(* Logix 5000 project; controller MV vendor 1 type 14 code 217 rev 31.11; software revision 31.00; part 32 of 53 *)
(* tags used below, declared in another part *)
   Alarm_Reset : BOOL;
   CWD : CHECKWORD_FLAGS;
   Default_Check_Time : DINT;
   FVHR12_1701 : PlantItem;   // Valve FVHR12_17/01
   FVHR12_1701_ALARM : ALARM_DIGITAL;
   FVHR12_1701_CL : ALIAS FOR RIO_Rack_2:13:I.Data.0;   // Valve FVHR12_17/01 Closed
   FVHR12_1701_DR : ALIAS FOR RIO_Rack_2:15:O.Data.0;   // Valve FVHR12_17/01 Drive
   FVHR12_1701_OP : ALIAS FOR RIO_Rack_2:13:I.Data.1;   // Valve FVHR12_17/01 Open
   FVHR12_1702 : PlantItem;   // Valve FVHR12_17/02
   FVHR12_1702_ALARM : ALARM_DIGITAL;
   FVHR12_1702_CL : ALIAS FOR RIO_Rack_2:13:I.Data.2;   // Valve FVHR12_17/02 Closed
   FVHR12_1702_DR : ALIAS FOR RIO_Rack_2:15:O.Data.1;   // Valve FVHR12_17/02 Drive
   FVHR12_1702_OP : ALIAS FOR RIO_Rack_2:13:I.Data.3;   // Valve FVHR12_17/02 Open
   FVHR12_1703 : PlantItem;   // Valve FVHR12_17/03
   FVHR12_1703_ALARM : ALARM_DIGITAL;
   FVHR12_1703_CL : ALIAS FOR RIO_Rack_2:13:I.Data.10;   // Valve FVHR12_17/03 Closed
   FVHR12_1703_DR : ALIAS FOR RIO_Rack_2:15:O.Data.5;   // Valve FVHR12_17/03 Drive
   FVHR12_1703_OP : ALIAS FOR RIO_Rack_2:13:I.Data.11;   // Valve FVHR12_17/03 Open
   FVHR18_2501 : PlantItem;   // Valve FVHR18_25/01
   FVHR18_2501_ALARM : ALARM_DIGITAL;
   FVHR18_2501_CL : ALIAS FOR RIO_Rack_2:13:I.Data.18;   // Valve FVHR18_25/01 Closed
   FVHR18_2501_DR : ALIAS FOR RIO_Rack_2:15:O.Data.9;   // Valve FVHR18_25/01 Drive
   FVHR18_2501_OP : ALIAS FOR RIO_Rack_2:13:I.Data.19;   // Valve FVHR18_25/01 Open
   FVHR18_2502 : PlantItem;   // Valve FVHR18_25/02
   FVHR18_2502_ALARM : ALARM_DIGITAL;
   FVHR18_2502_CL : ALIAS FOR RIO_Rack_2:13:I.Data.20;   // Valve FVHR18_25/02 Closed
   FVHR18_2502_DR : ALIAS FOR RIO_Rack_2:15:O.Data.10;   // Valve FVHR18_25/02 Drive
   FVHR18_2502_OP : ALIAS FOR RIO_Rack_2:13:I.Data.21;   // Valve FVHR18_25/02 Open
   FVHR18_2503 : PlantItem;   // Valve FVHR18_25/03
   FVHR18_2503_ALARM : ALARM_DIGITAL;
   FVHR18_2503_CL : ALIAS FOR RIO_Rack_2:13:I.Data.22;   // Valve FVHR18_25/03 Closed
   FVHR18_2503_DR : ALIAS FOR RIO_Rack_2:15:O.Data.11;   // Valve FVHR18_25/03 Drive
   FVHR18_2503_OP : ALIAS FOR RIO_Rack_2:13:I.Data.23;   // Valve FVHR18_25/03 Open
   FVHR18_2504 : PlantItem;   // Valve FVHR18_25/04
   FVHR18_2504_ALARM : ALARM_DIGITAL;
   FVHR18_2504_CL : ALIAS FOR RIO_Rack_2:13:I.Data.24;   // Valve FVHR18_25/04 Closed
   FVHR18_2504_DR : ALIAS FOR RIO_Rack_2:15:O.Data.12;   // Valve FVHR18_25/04 Drive
   FVHR18_2504_OP : ALIAS FOR RIO_Rack_2:13:I.Data.25;   // Valve FVHR18_25/04 Open
   FVHR18_2505 : PlantItem;   // Valve FVHR18_25/05
   FVHR18_2505_ALARM : ALARM_DIGITAL;
   FVHR18_2505_CL : ALIAS FOR RIO_Rack_2:13:I.Data.26;   // Valve FVHR18_25/05 Closed
   FVHR18_2505_DR : ALIAS FOR RIO_Rack_2:15:O.Data.13;   // Valve FVHR18_25/05 Drive
   FVHR18_2505_OP : ALIAS FOR RIO_Rack_2:13:I.Data.27;   // Valve FVHR18_25/05 Open
   FVHR18_2506 : PlantItem;   // Valve FVHR18_25/06
   FVHR18_2506_ALARM : ALARM_DIGITAL;
   FVHR18_2506_CL : ALIAS FOR RIO_Rack_2:13:I.Data.28;   // Valve FVHR18_25/06 Closed
   FVHR18_2506_DR : ALIAS FOR RIO_Rack_2:15:O.Data.14;   // Valve FVHR18_25/06 Drive
   FVHR18_2506_OP : ALIAS FOR RIO_Rack_2:13:I.Data.29;   // Valve FVHR18_25/06 Open
   FVHR1_1101 : PlantItem;   // Valve FVHR1_11/01
   FVHR1_1101_ALARM : ALARM_DIGITAL;
   FVHR1_1101_CL : ALIAS FOR RIO_Rack_2:13:I.Data.4;   // Valve FVHR1_11/01 Closed
   FVHR1_1101_DR : ALIAS FOR RIO_Rack_2:15:O.Data.2;   // Valve FVHR1_11/01 Drive
   FVHR1_1101_OP : ALIAS FOR RIO_Rack_2:13:I.Data.5;   // Valve FVHR1_11/01 Open
   FVHR1_1102 : PlantItem;   // Valve FVHR1_11/02
   FVHR1_1102_ALARM : ALARM_DIGITAL;
   FVHR1_1102_CL : ALIAS FOR RIO_Rack_2:13:I.Data.6;   // Valve FVHR1_11/02 Closed
   FVHR1_1102_DR : ALIAS FOR RIO_Rack_2:15:O.Data.3;   // Valve FVHR1_11/02 Drive
   FVHR1_1102_OP : ALIAS FOR RIO_Rack_2:13:I.Data.7;   // Valve FVHR1_11/02 Open
   FVHR1_1103 : PlantItem;   // Valve FVHR1_11/03
   FVHR1_1103_ALARM : ALARM_DIGITAL;
   FVHR1_1103_CL : ALIAS FOR RIO_Rack_2:13:I.Data.8;   // Valve FVHR1_11/03 Closed
   FVHR1_1103_DR : ALIAS FOR RIO_Rack_2:15:O.Data.4;   // Valve FVHR1_11/03 Drive
   FVHR1_1103_OP : ALIAS FOR RIO_Rack_2:13:I.Data.9;   // Valve FVHR1_11/03 Open
   FVHR1_1701 : PlantItem;   // Valve FVHR1_17/01
   FVHR1_1701_ALARM : ALARM_DIGITAL;
   FVHR1_1701_CL : ALIAS FOR RIO_Rack_2:13:I.Data.16;   // Valve FVHR1_17/01 Closed
   FVHR1_1701_DR : ALIAS FOR RIO_Rack_2:15:O.Data.8;   // Valve FVHR1_17/01 Drive
   FVHR1_1701_OP : ALIAS FOR RIO_Rack_2:13:I.Data.17;   // Valve FVHR1_17/01 Open
   FVHR26_3101 : PlantItem;   // Valve FVHR26_31/01
   FVHR26_3101_ALARM : ALARM_DIGITAL;
   FVHR26_3101_CL : ALIAS FOR RIO_Rack_2:14:I.Data.2;   // Valve FVHR26_31/01 Closed
   FVHR26_3101_DR : ALIAS FOR RIO_Rack_2:15:O.Data.17;   // Valve FVHR26_31/01 Drive
   FVHR26_3101_OP : ALIAS FOR RIO_Rack_2:14:I.Data.3;   // Valve FVHR26_31/01 Open
   IGI_TestBit : BOOL;
   Item_Faults_Are_Latched : BOOL;
   Item_Simulation_Flag : BOOL;
   MC_CIP_AV01 : PlantItem;   // CIP_AV01
   MC_CIP_AV01_ALARM : ALARM_DIGITAL;
   MC_CIP_AV01_C : ALIAS FOR RIO_Rack_2:9:I.Data.23;
   MC_CIP_AV01_DR : ALIAS FOR CIP_AV01_DUMMY_DR;
   MC_CIP_AV01_O : ALIAS FOR RIO_Rack_2:9:I.Data.19;
   MC_CIP_AV02 : PlantItem;   // CIP_AV02
   MC_CIP_AV02_ALARM : ALARM_DIGITAL;
   MC_CIP_AV02_C : ALIAS FOR RIO_Rack_2:9:I.Data.28;
   MC_CIP_AV02_DR : ALIAS FOR RIO_Rack_2:8:O.Data.27;   // Used As Output Share Item Rung 20
   MC_CIP_AV02_O : ALIAS FOR RIO_Rack_2:9:I.Data.24;
   MC_CIP_AV05 : PlantItem;   // CIP_AV05
   MC_CIP_AV05_ALARM : ALARM_DIGITAL;
   MC_CIP_AV05_C : ALIAS FOR RIO_Rack_2:9:I.Data.29;
   MC_CIP_AV05_DR : ALIAS FOR CIP_AV05_DUMMY_DR;
   MC_CIP_AV05_O : ALIAS FOR RIO_Rack_2:9:I.Data.25;
   MC_CIP_AV06 : PlantItem;   // CIP_AV06
   MC_CIP_AV06_ALARM : ALARM_DIGITAL;
   MC_CIP_AV06_C : ALIAS FOR RIO_Rack_2:9:I.Data.30;
   MC_CIP_AV06_DR : ALIAS FOR RIO_Rack_2:8:O.Data.28;
   MC_CIP_AV06_O : ALIAS FOR RIO_Rack_2:9:I.Data.26;
   MC_CIP_AV07 : PlantItem;   // CIP_AV07
   MC_CIP_AV07_ALARM : ALARM_DIGITAL;
   MC_CIP_AV07_C : ALIAS FOR RIO_Rack_2:9:I.Data.31;
   MC_CIP_AV07_DR : ALIAS FOR CIP_AV07_DUMMY_DR;
   MC_CIP_AV07_O : ALIAS FOR RIO_Rack_2:9:I.Data.27;
   MC_CIP_AV08 : PlantItem;   // CIP_AV08
   MC_CIP_AV08_ALARM : ALARM_DIGITAL;
   MC_CIP_AV08_C : ALIAS FOR RIO_Rack_2:11:I.Data.20;
   MC_CIP_AV08_DR : ALIAS FOR RIO_Rack_2:8:O.Data.29;
   MC_CIP_AV08_O : ALIAS FOR RIO_Rack_2:11:I.Data.24;
   MC_CIP_AV09 : PlantItem;   // CIP_AV09
   MC_CIP_AV09_ALARM : ALARM_DIGITAL;
   MC_CIP_AV09_C : ALIAS FOR RIO_Rack_2:11:I.Data.21;
   MC_CIP_AV09_DR : ALIAS FOR CIP_AV09_DUMMY_DR;
   MC_CIP_AV09_O : ALIAS FOR RIO_Rack_2:11:I.Data.25;
   MC_CIP_AV10 : PlantItem;   // CIP_AV10
   MC_CIP_AV10_ALARM : ALARM_DIGITAL;
   MC_CIP_AV10_C : ALIAS FOR RIO_Rack_2:11:I.Data.22;
   MC_CIP_AV10_DR : ALIAS FOR RIO_Rack_2:8:O.Data.30;
   MC_CIP_AV10_O : ALIAS FOR RIO_Rack_2:11:I.Data.26;
   MC_CIP_RV : PlantItem;   // CIP_RV
   MC_CIP_RV_ALARM : ALARM_DIGITAL;
   MC_CIP_RV_C : ALIAS FOR RIO_Rack_2:9:I.Data.21;
   MC_CIP_RV_DR : ALIAS FOR RIO_Rack_2:8:O.Data.26;
   MC_CIP_RV_O : ALIAS FOR RIO_Rack_2:9:I.Data.17;
   MC_R3R_DR : PlantItem;   // R3R_DR
   MC_R3R_DR_ALARM : ALARM_DIGITAL;
   MC_R3R_DR_C : ALIAS FOR RIO_Rack_2:9:I.Data.20;
   MC_R3R_DR_DR : ALIAS FOR RIO_Rack_2:8:O.Data.24;
   MC_R3R_DR_O : ALIAS FOR RIO_Rack_2:9:I.Data.16;
   One_Second_One_Scan : ALIAS FOR One_Second_1_scan;
(* MC_Common, continued *)

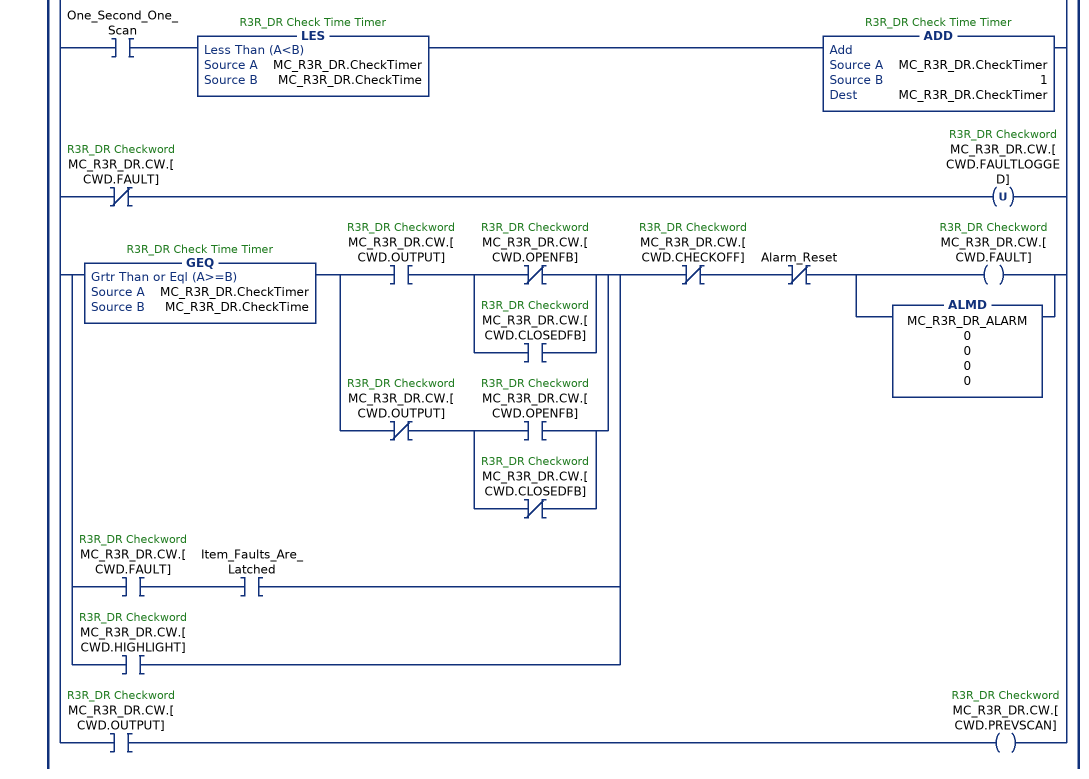
   [picture p709: MC_Common/MC_Valves rungs 55-55]
   55: [NEQ(MC_R3R_DR.DriveBits,0) OTE(MC_R3R_DR.CW.[CWD.AUTODRV]) ,[XIC(MC_R3R_DR.CW.[CWD.AUTODRV]) XIO(MC_R3R_DR.CW.[CWD.MANUAL]) ,XIC(MC_R3R_DR.CW.[CWD.MANDRV]) XIC(MC_R3R_DR.CW.[CWD.MANUAL]) ] OTE(MC_R3R_DR.CW.[CWD.OUTPUT]) ,XIC(MC_R3R_DR.CW.[CWD.OUTPUT]) OTE(MC_R3R_DR_DR) ,XIC(S:FS) [OTU(MC_R3R_DR.CW.[CWD.MANUAL]) ,LEQ(MC_R3R_DR.CheckTime,0) MOV(Default_Check_Time,MC_R3R_DR.CheckTime) ] ,[[XIC(MC_R3R_DR_O) XIO(Item_Simulation_Flag) ,XIC(Item_Simulation_Flag) XIC(MC_R3R_DR.CW.[CWD.OUTPUT]) XIO(MC_R3R_DR.CW.[CWD.SIMFAIL]) ] OTE(MC_R3R_DR.CW.[CWD.OPENFB]) ,[XIC(MC_R3R_DR_C) XIO(Item_Simulation_Flag) ,XIC(Item_Simulation_Flag) XIO(MC_R3R_DR.CW.[CWD.OUTPUT]) XIO(MC_R3R_DR.CW.[CWD.SIMFAIL]) ] OTE(MC_R3R_DR.CW.[CWD.CLOSEDFB]) ] ,[XIC(MC_R3R_DR.CW.[CWD.OUTPUT]) XIO(MC_R3R_DR.CW.[CWD.PREVSCAN]) ,XIO(MC_R3R_DR.CW.[CWD.OUTPUT]) XIC(MC_R3R_DR.CW.[CWD.PREVSCAN]) ] CLR(MC_R3R_DR.CheckTimer) ,XIC(One_Second_One_Scan) LES(MC_R3R_DR.CheckTimer,MC_R3R_DR.CheckTime) ADD(MC_R3R_DR.CheckTimer,1,MC_R3R_DR.CheckTimer) ,XIO(MC_R3R_DR.CW.[CWD.FAULT]) OTU(MC_R3R_DR.CW.[CWD.FAULTLOGGED]) ,[GEQ(MC_R3R_DR.CheckTimer,MC_R3R_DR.CheckTime) [XIC(MC_R3R_DR.CW.[CWD.OUTPUT]) [XIO(MC_R3R_DR.CW.[CWD.OPENFB]) ,XIC(MC_R3R_DR.CW.[CWD.CLOSEDFB]) ] ,XIO(MC_R3R_DR.CW.[CWD.OUTPUT]) [XIC(MC_R3R_DR.CW.[CWD.OPENFB]) ,XIO(MC_R3R_DR.CW.[CWD.CLOSEDFB]) ] ] ,XIC(MC_R3R_DR.CW.[CWD.FAULT]) XIC(Item_Faults_Are_Latched) ,XIC(MC_R3R_DR.CW.[CWD.HIGHLIGHT]) ] XIO(MC_R3R_DR.CW.[CWD.CHECKOFF]) XIO(Alarm_Reset) [OTE(MC_R3R_DR.CW.[CWD.FAULT]) ,ALMD(MC_R3R_DR_ALARM,0,0,0,0) ] ,XIC(MC_R3R_DR.CW.[CWD.OUTPUT]) OTE(MC_R3R_DR.CW.[CWD.PREVSCAN]) ];
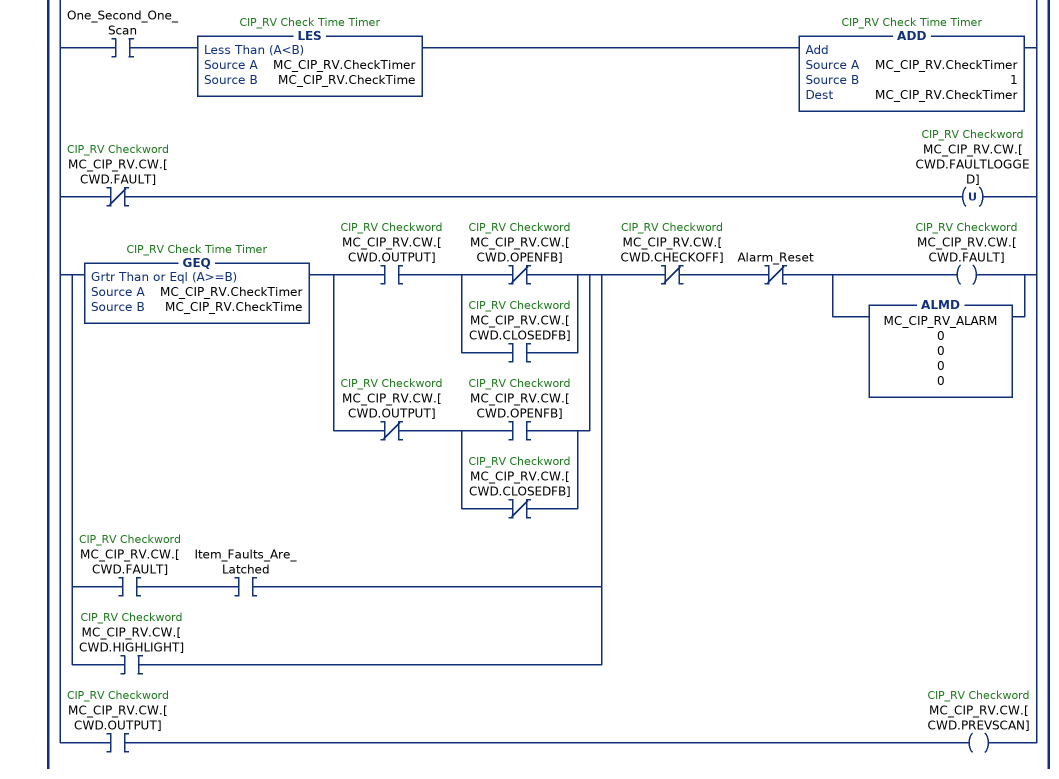
   56: [NEQ(MC_CIP_RV.DriveBits,0) OTE(MC_CIP_RV.CW.[CWD.AUTODRV]) ,[XIC(MC_CIP_RV.CW.[CWD.AUTODRV]) XIO(MC_CIP_RV.CW.[CWD.MANUAL]) ,XIC(MC_CIP_RV.CW.[CWD.MANDRV]) XIC(MC_CIP_RV.CW.[CWD.MANUAL]) ] OTE(MC_CIP_RV.CW.[CWD.OUTPUT]) ,XIC(MC_CIP_RV.CW.[CWD.OUTPUT]) OTE(MC_CIP_RV_DR) ,XIC(S:FS) [OTU(MC_CIP_RV.CW.[CWD.MANUAL]) ,LEQ(MC_CIP_RV.CheckTime,0) MOV(Default_Check_Time,MC_CIP_RV.CheckTime) ] ,[[XIC(MC_CIP_RV_O) XIO(Item_Simulation_Flag) ,XIC(Item_Simulation_Flag) XIC(MC_CIP_RV.CW.[CWD.OUTPUT]) XIO(MC_CIP_RV.CW.[CWD.SIMFAIL]) ] OTE(MC_CIP_RV.CW.[CWD.OPENFB]) ,[XIC(MC_CIP_RV_C) XIO(Item_Simulation_Flag) ,XIC(Item_Simulation_Flag) XIO(MC_CIP_RV.CW.[CWD.OUTPUT]) XIO(MC_CIP_RV.CW.[CWD.SIMFAIL]) ] OTE(MC_CIP_RV.CW.[CWD.CLOSEDFB]) ] ,[XIC(MC_CIP_RV.CW.[CWD.OUTPUT]) XIO(MC_CIP_RV.CW.[CWD.PREVSCAN]) ,XIO(MC_CIP_RV.CW.[CWD.OUTPUT]) XIC(MC_CIP_RV.CW.[CWD.PREVSCAN]) ] CLR(MC_CIP_RV.CheckTimer) ,XIC(One_Second_One_Scan) LES(MC_CIP_RV.CheckTimer,MC_CIP_RV.CheckTime) ADD(MC_CIP_RV.CheckTimer,1,MC_CIP_RV.CheckTimer) ,XIO(MC_CIP_RV.CW.[CWD.FAULT]) OTU(MC_CIP_RV.CW.[CWD.FAULTLOGGED]) ,[GEQ(MC_CIP_RV.CheckTimer,MC_CIP_RV.CheckTime) [XIC(MC_CIP_RV.CW.[CWD.OUTPUT]) [XIO(MC_CIP_RV.CW.[CWD.OPENFB]) ,XIC(MC_CIP_RV.CW.[CWD.CLOSEDFB]) ] ,XIO(MC_CIP_RV.CW.[CWD.OUTPUT]) [XIC(MC_CIP_RV.CW.[CWD.OPENFB]) ,XIO(MC_CIP_RV.CW.[CWD.CLOSEDFB]) ] ] ,XIC(MC_CIP_RV.CW.[CWD.FAULT]) XIC(Item_Faults_Are_Latched) ,XIC(MC_CIP_RV.CW.[CWD.HIGHLIGHT]) ] XIO(MC_CIP_RV.CW.[CWD.CHECKOFF]) XIO(Alarm_Reset) [OTE(MC_CIP_RV.CW.[CWD.FAULT]) ,ALMD(MC_CIP_RV_ALARM,0,0,0,0) ] ,XIC(MC_CIP_RV.CW.[CWD.OUTPUT]) OTE(MC_CIP_RV.CW.[CWD.PREVSCAN]) ];
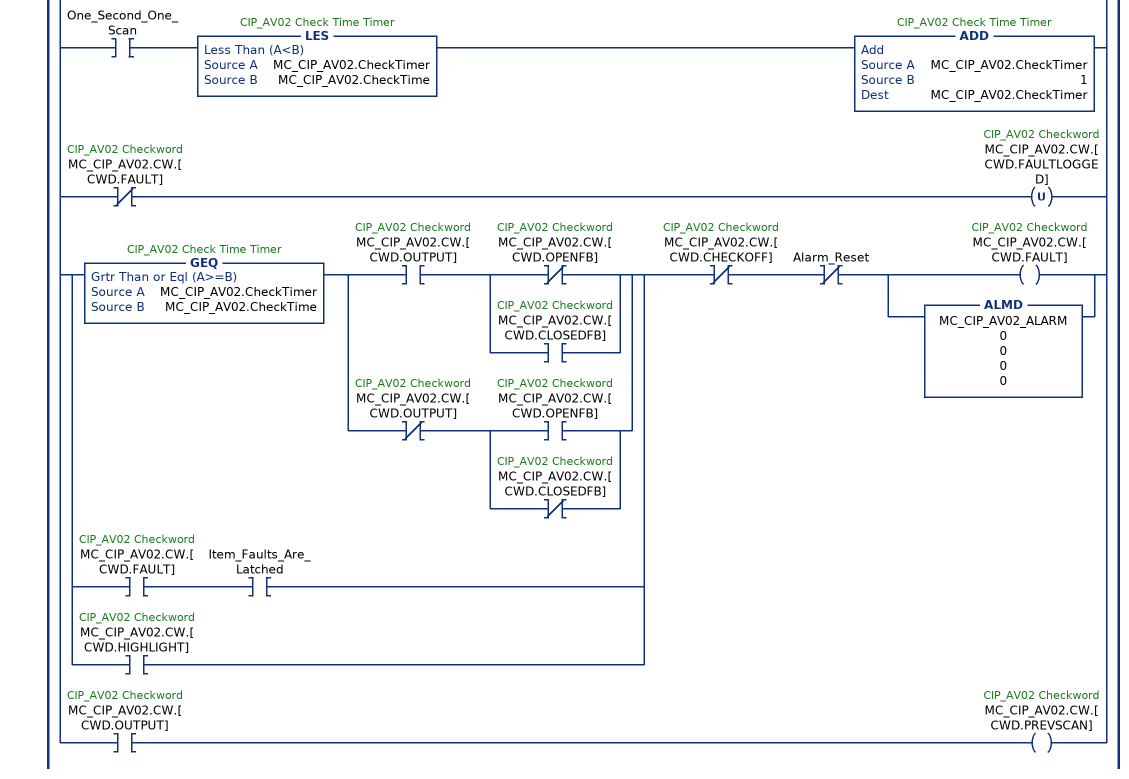
   57: [NEQ(MC_CIP_AV02.DriveBits,0) OTE(MC_CIP_AV02.CW.[CWD.AUTODRV]) ,[XIC(MC_CIP_AV02.CW.[CWD.AUTODRV]) XIO(MC_CIP_AV02.CW.[CWD.MANUAL]) ,XIC(MC_CIP_AV02.CW.[CWD.MANDRV]) XIC(MC_CIP_AV02.CW.[CWD.MANUAL]) ] OTE(MC_CIP_AV02.CW.[CWD.OUTPUT]) ,XIC(MC_CIP_AV02.CW.[CWD.OUTPUT]) OTE(MC_CIP_AV02_DR) ,XIC(S:FS) [OTU(MC_CIP_AV02.CW.[CWD.MANUAL]) ,LEQ(MC_CIP_AV02.CheckTime,0) MOV(Default_Check_Time,MC_CIP_AV02.CheckTime) ] ,[[XIC(MC_CIP_AV02_O) XIO(Item_Simulation_Flag) ,XIC(Item_Simulation_Flag) XIC(MC_CIP_AV02.CW.[CWD.OUTPUT]) XIO(MC_CIP_AV02.CW.[CWD.SIMFAIL]) ] OTE(MC_CIP_AV02.CW.[CWD.OPENFB]) ,[XIC(MC_CIP_AV02_C) XIO(Item_Simulation_Flag) ,XIC(Item_Simulation_Flag) XIO(MC_CIP_AV02.CW.[CWD.OUTPUT]) XIO(MC_CIP_AV02.CW.[CWD.SIMFAIL]) ] OTE(MC_CIP_AV02.CW.[CWD.CLOSEDFB]) ] ,[XIC(MC_CIP_AV02.CW.[CWD.OUTPUT]) XIO(MC_CIP_AV02.CW.[CWD.PREVSCAN]) ,XIO(MC_CIP_AV02.CW.[CWD.OUTPUT]) XIC(MC_CIP_AV02.CW.[CWD.PREVSCAN]) ] CLR(MC_CIP_AV02.CheckTimer) ,XIC(One_Second_One_Scan) LES(MC_CIP_AV02.CheckTimer,MC_CIP_AV02.CheckTime) ADD(MC_CIP_AV02.CheckTimer,1,MC_CIP_AV02.CheckTimer) ,XIO(MC_CIP_AV02.CW.[CWD.FAULT]) OTU(MC_CIP_AV02.CW.[CWD.FAULTLOGGED]) ,[GEQ(MC_CIP_AV02.CheckTimer,MC_CIP_AV02.CheckTime) [XIC(MC_CIP_AV02.CW.[CWD.OUTPUT]) [XIO(MC_CIP_AV02.CW.[CWD.OPENFB]) ,XIC(MC_CIP_AV02.CW.[CWD.CLOSEDFB]) ] ,XIO(MC_CIP_AV02.CW.[CWD.OUTPUT]) [XIC(MC_CIP_AV02.CW.[CWD.OPENFB]) ,XIO(MC_CIP_AV02.CW.[CWD.CLOSEDFB]) ] ] ,XIC(MC_CIP_AV02.CW.[CWD.FAULT]) XIC(Item_Faults_Are_Latched) ,XIC(MC_CIP_AV02.CW.[CWD.HIGHLIGHT]) ] XIO(MC_CIP_AV02.CW.[CWD.CHECKOFF]) XIO(Alarm_Reset) [OTE(MC_CIP_AV02.CW.[CWD.FAULT]) ,ALMD(MC_CIP_AV02_ALARM,0,0,0,0) ] ,XIC(MC_CIP_AV02.CW.[CWD.OUTPUT]) OTE(MC_CIP_AV02.CW.[CWD.PREVSCAN]) ];
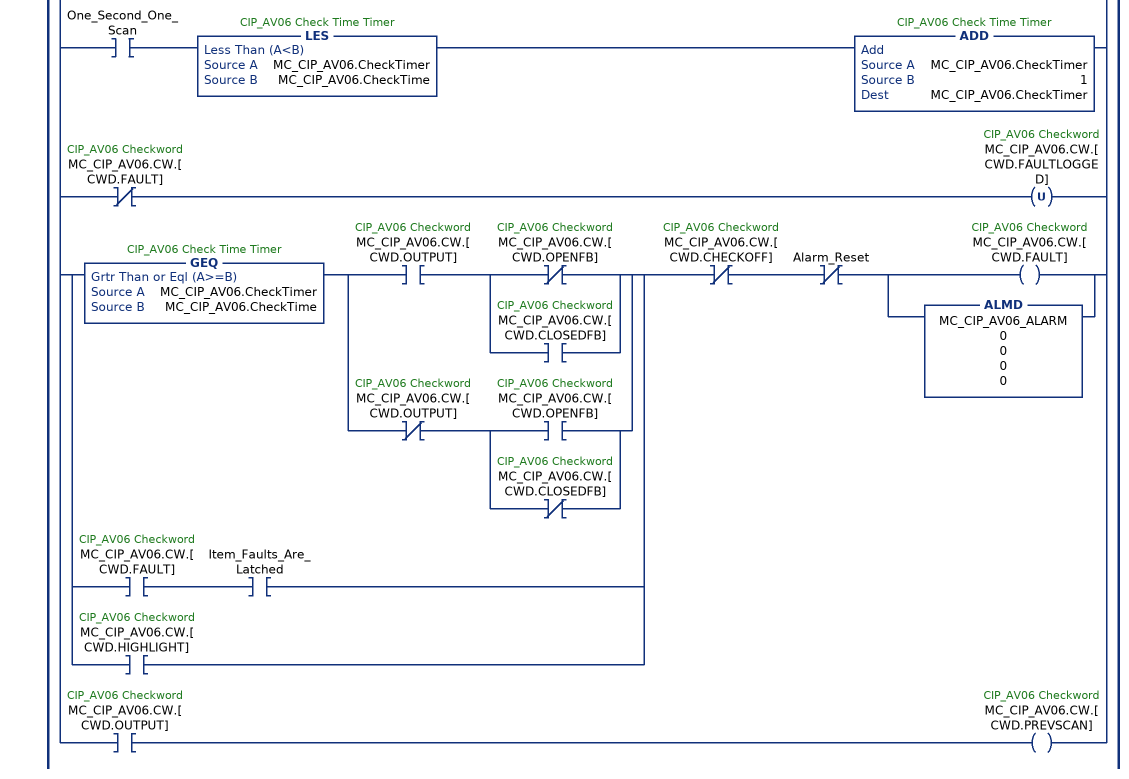
   58: [NEQ(MC_CIP_AV06.DriveBits,0) OTE(MC_CIP_AV06.CW.[CWD.AUTODRV]) ,[XIC(MC_CIP_AV06.CW.[CWD.AUTODRV]) XIO(MC_CIP_AV06.CW.[CWD.MANUAL]) ,XIC(MC_CIP_AV06.CW.[CWD.MANDRV]) XIC(MC_CIP_AV06.CW.[CWD.MANUAL]) ] OTE(MC_CIP_AV06.CW.[CWD.OUTPUT]) ,XIC(MC_CIP_AV06.CW.[CWD.OUTPUT]) OTE(MC_CIP_AV06_DR) ,XIC(S:FS) [OTU(MC_CIP_AV06.CW.[CWD.MANUAL]) ,LEQ(MC_CIP_AV06.CheckTime,0) MOV(Default_Check_Time,MC_CIP_AV06.CheckTime) ] ,[[XIC(MC_CIP_AV06_O) XIO(Item_Simulation_Flag) ,XIC(Item_Simulation_Flag) XIC(MC_CIP_AV06.CW.[CWD.OUTPUT]) XIO(MC_CIP_AV06.CW.[CWD.SIMFAIL]) ] OTE(MC_CIP_AV06.CW.[CWD.OPENFB]) ,[XIC(MC_CIP_AV06_C) XIO(Item_Simulation_Flag) ,XIC(Item_Simulation_Flag) XIO(MC_CIP_AV06.CW.[CWD.OUTPUT]) XIO(MC_CIP_AV06.CW.[CWD.SIMFAIL]) ] OTE(MC_CIP_AV06.CW.[CWD.CLOSEDFB]) ] ,[XIC(MC_CIP_AV06.CW.[CWD.OUTPUT]) XIO(MC_CIP_AV06.CW.[CWD.PREVSCAN]) ,XIO(MC_CIP_AV06.CW.[CWD.OUTPUT]) XIC(MC_CIP_AV06.CW.[CWD.PREVSCAN]) ] CLR(MC_CIP_AV06.CheckTimer) ,XIC(One_Second_One_Scan) LES(MC_CIP_AV06.CheckTimer,MC_CIP_AV06.CheckTime) ADD(MC_CIP_AV06.CheckTimer,1,MC_CIP_AV06.CheckTimer) ,XIO(MC_CIP_AV06.CW.[CWD.FAULT]) OTU(MC_CIP_AV06.CW.[CWD.FAULTLOGGED]) ,[GEQ(MC_CIP_AV06.CheckTimer,MC_CIP_AV06.CheckTime) [XIC(MC_CIP_AV06.CW.[CWD.OUTPUT]) [XIO(MC_CIP_AV06.CW.[CWD.OPENFB]) ,XIC(MC_CIP_AV06.CW.[CWD.CLOSEDFB]) ] ,XIO(MC_CIP_AV06.CW.[CWD.OUTPUT]) [XIC(MC_CIP_AV06.CW.[CWD.OPENFB]) ,XIO(MC_CIP_AV06.CW.[CWD.CLOSEDFB]) ] ] ,XIC(MC_CIP_AV06.CW.[CWD.FAULT]) XIC(Item_Faults_Are_Latched) ,XIC(MC_CIP_AV06.CW.[CWD.HIGHLIGHT]) ] XIO(MC_CIP_AV06.CW.[CWD.CHECKOFF]) XIO(Alarm_Reset) [OTE(MC_CIP_AV06.CW.[CWD.FAULT]) ,ALMD(MC_CIP_AV06_ALARM,0,0,0,0) ] ,XIC(MC_CIP_AV06.CW.[CWD.OUTPUT]) OTE(MC_CIP_AV06.CW.[CWD.PREVSCAN]) ];
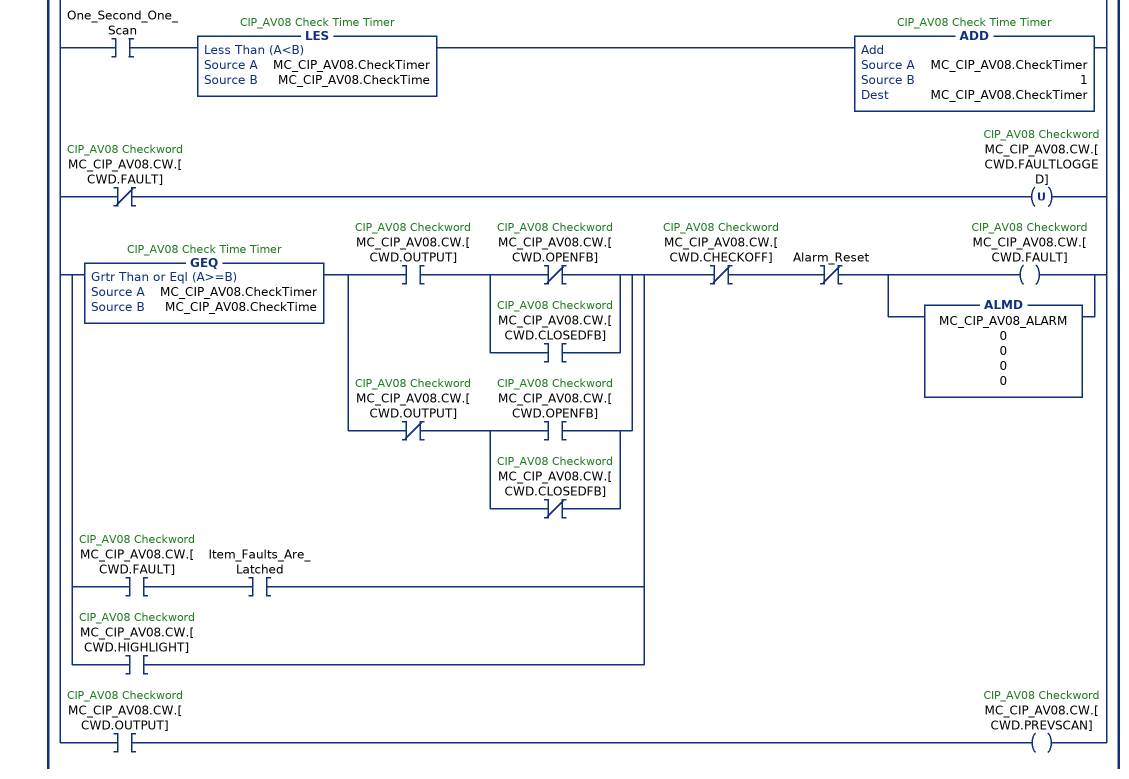
   59: [NEQ(MC_CIP_AV08.DriveBits,0) OTE(MC_CIP_AV08.CW.[CWD.AUTODRV]) ,[XIC(MC_CIP_AV08.CW.[CWD.AUTODRV]) XIO(MC_CIP_AV08.CW.[CWD.MANUAL]) ,XIC(MC_CIP_AV08.CW.[CWD.MANDRV]) XIC(MC_CIP_AV08.CW.[CWD.MANUAL]) ] OTE(MC_CIP_AV08.CW.[CWD.OUTPUT]) ,XIC(MC_CIP_AV08.CW.[CWD.OUTPUT]) OTE(MC_CIP_AV08_DR) ,XIC(S:FS) [OTU(MC_CIP_AV08.CW.[CWD.MANUAL]) ,LEQ(MC_CIP_AV08.CheckTime,0) MOV(Default_Check_Time,MC_CIP_AV08.CheckTime) ] ,[[XIC(MC_CIP_AV08_O) XIO(Item_Simulation_Flag) ,XIC(Item_Simulation_Flag) XIC(MC_CIP_AV08.CW.[CWD.OUTPUT]) XIO(MC_CIP_AV08.CW.[CWD.SIMFAIL]) ] OTE(MC_CIP_AV08.CW.[CWD.OPENFB]) ,[XIC(MC_CIP_AV08_C) XIO(Item_Simulation_Flag) ,XIC(Item_Simulation_Flag) XIO(MC_CIP_AV08.CW.[CWD.OUTPUT]) XIO(MC_CIP_AV08.CW.[CWD.SIMFAIL]) ] OTE(MC_CIP_AV08.CW.[CWD.CLOSEDFB]) ] ,[XIC(MC_CIP_AV08.CW.[CWD.OUTPUT]) XIO(MC_CIP_AV08.CW.[CWD.PREVSCAN]) ,XIO(MC_CIP_AV08.CW.[CWD.OUTPUT]) XIC(MC_CIP_AV08.CW.[CWD.PREVSCAN]) ] CLR(MC_CIP_AV08.CheckTimer) ,XIC(One_Second_One_Scan) LES(MC_CIP_AV08.CheckTimer,MC_CIP_AV08.CheckTime) ADD(MC_CIP_AV08.CheckTimer,1,MC_CIP_AV08.CheckTimer) ,XIO(MC_CIP_AV08.CW.[CWD.FAULT]) OTU(MC_CIP_AV08.CW.[CWD.FAULTLOGGED]) ,[GEQ(MC_CIP_AV08.CheckTimer,MC_CIP_AV08.CheckTime) [XIC(MC_CIP_AV08.CW.[CWD.OUTPUT]) [XIO(MC_CIP_AV08.CW.[CWD.OPENFB]) ,XIC(MC_CIP_AV08.CW.[CWD.CLOSEDFB]) ] ,XIO(MC_CIP_AV08.CW.[CWD.OUTPUT]) [XIC(MC_CIP_AV08.CW.[CWD.OPENFB]) ,XIO(MC_CIP_AV08.CW.[CWD.CLOSEDFB]) ] ] ,XIC(MC_CIP_AV08.CW.[CWD.FAULT]) XIC(Item_Faults_Are_Latched) ,XIC(MC_CIP_AV08.CW.[CWD.HIGHLIGHT]) ] XIO(MC_CIP_AV08.CW.[CWD.CHECKOFF]) XIO(Alarm_Reset) [OTE(MC_CIP_AV08.CW.[CWD.FAULT]) ,ALMD(MC_CIP_AV08_ALARM,0,0,0,0) ] ,XIC(MC_CIP_AV08.CW.[CWD.OUTPUT]) OTE(MC_CIP_AV08.CW.[CWD.PREVSCAN]) ];
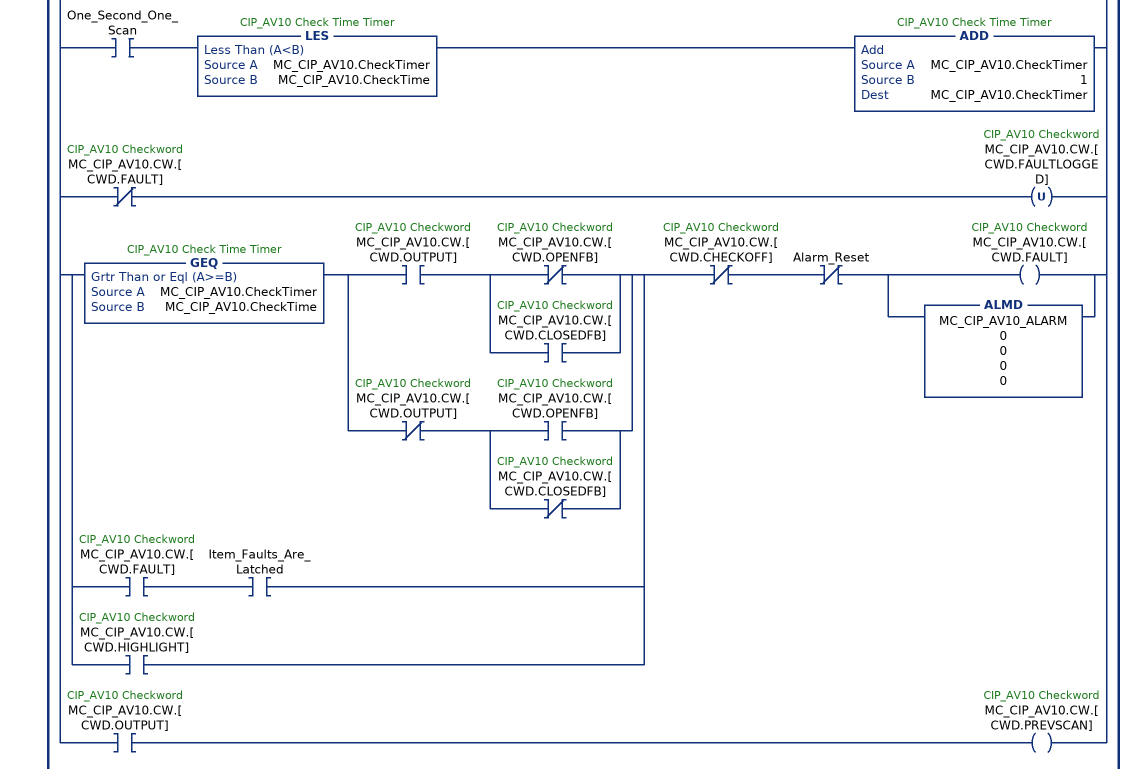
   60: [NEQ(MC_CIP_AV10.DriveBits,0) OTE(MC_CIP_AV10.CW.[CWD.AUTODRV]) ,[XIC(MC_CIP_AV10.CW.[CWD.AUTODRV]) XIO(MC_CIP_AV10.CW.[CWD.MANUAL]) ,XIC(MC_CIP_AV10.CW.[CWD.MANDRV]) XIC(MC_CIP_AV10.CW.[CWD.MANUAL]) ] OTE(MC_CIP_AV10.CW.[CWD.OUTPUT]) ,XIC(MC_CIP_AV10.CW.[CWD.OUTPUT]) OTE(MC_CIP_AV10_DR) ,XIC(S:FS) [OTU(MC_CIP_AV10.CW.[CWD.MANUAL]) ,LEQ(MC_CIP_AV10.CheckTime,0) MOV(Default_Check_Time,MC_CIP_AV10.CheckTime) ] ,[[XIC(MC_CIP_AV10_O) XIO(Item_Simulation_Flag) ,XIC(Item_Simulation_Flag) XIC(MC_CIP_AV10.CW.[CWD.OUTPUT]) XIO(MC_CIP_AV10.CW.[CWD.SIMFAIL]) ] OTE(MC_CIP_AV10.CW.[CWD.OPENFB]) ,[XIC(MC_CIP_AV10_C) XIO(Item_Simulation_Flag) ,XIC(Item_Simulation_Flag) XIO(MC_CIP_AV10.CW.[CWD.OUTPUT]) XIO(MC_CIP_AV10.CW.[CWD.SIMFAIL]) ] OTE(MC_CIP_AV10.CW.[CWD.CLOSEDFB]) ] ,[XIC(MC_CIP_AV10.CW.[CWD.OUTPUT]) XIO(MC_CIP_AV10.CW.[CWD.PREVSCAN]) ,XIO(MC_CIP_AV10.CW.[CWD.OUTPUT]) XIC(MC_CIP_AV10.CW.[CWD.PREVSCAN]) ] CLR(MC_CIP_AV10.CheckTimer) ,XIC(One_Second_One_Scan) LES(MC_CIP_AV10.CheckTimer,MC_CIP_AV10.CheckTime) ADD(MC_CIP_AV10.CheckTimer,1,MC_CIP_AV10.CheckTimer) ,XIO(MC_CIP_AV10.CW.[CWD.FAULT]) OTU(MC_CIP_AV10.CW.[CWD.FAULTLOGGED]) ,[GEQ(MC_CIP_AV10.CheckTimer,MC_CIP_AV10.CheckTime) [XIC(MC_CIP_AV10.CW.[CWD.OUTPUT]) [XIO(MC_CIP_AV10.CW.[CWD.OPENFB]) ,XIC(MC_CIP_AV10.CW.[CWD.CLOSEDFB]) ] ,XIO(MC_CIP_AV10.CW.[CWD.OUTPUT]) [XIC(MC_CIP_AV10.CW.[CWD.OPENFB]) ,XIO(MC_CIP_AV10.CW.[CWD.CLOSEDFB]) ] ] ,XIC(MC_CIP_AV10.CW.[CWD.FAULT]) XIC(Item_Faults_Are_Latched) ,XIC(MC_CIP_AV10.CW.[CWD.HIGHLIGHT]) ] XIO(MC_CIP_AV10.CW.[CWD.CHECKOFF]) XIO(Alarm_Reset) [OTE(MC_CIP_AV10.CW.[CWD.FAULT]) ,ALMD(MC_CIP_AV10_ALARM,0,0,0,0) ] ,XIC(MC_CIP_AV10.CW.[CWD.OUTPUT]) OTE(MC_CIP_AV10.CW.[CWD.PREVSCAN]) ];
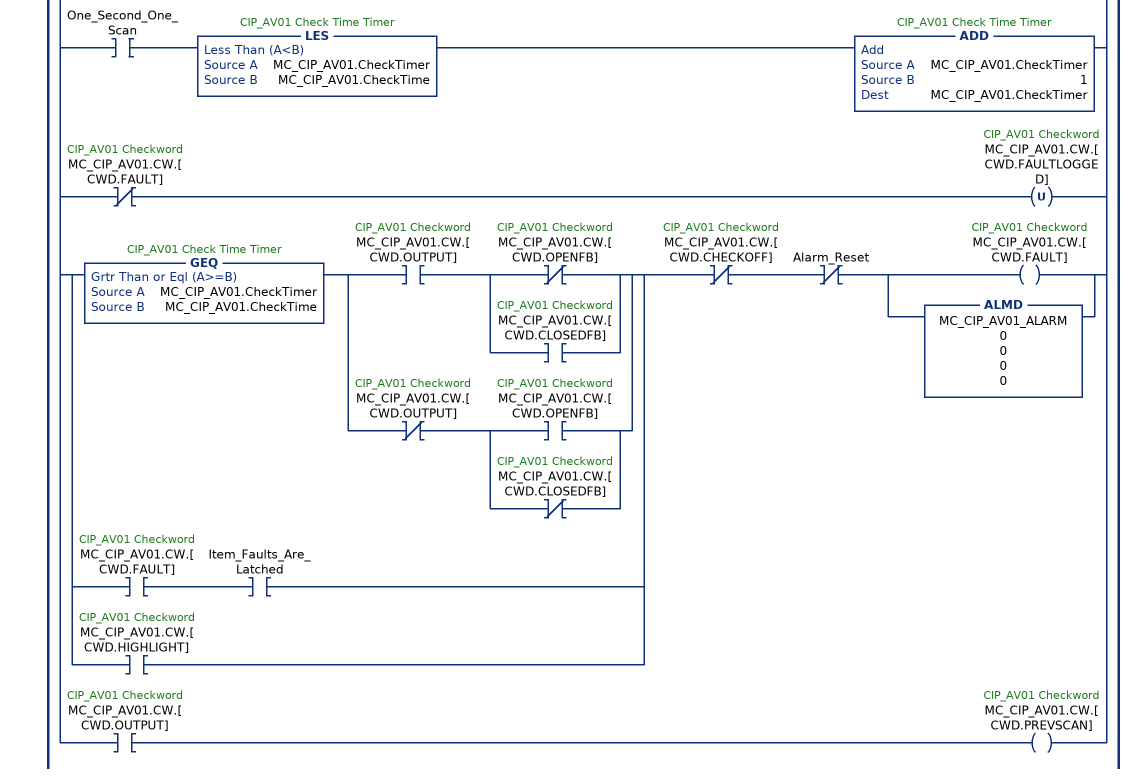
   61: [NEQ(MC_CIP_AV01.DriveBits,0) OTE(MC_CIP_AV01.CW.[CWD.AUTODRV]) ,[XIC(MC_CIP_AV01.CW.[CWD.AUTODRV]) XIO(MC_CIP_AV01.CW.[CWD.MANUAL]) ,XIC(MC_CIP_AV01.CW.[CWD.MANDRV]) XIC(MC_CIP_AV01.CW.[CWD.MANUAL]) ] OTE(MC_CIP_AV01.CW.[CWD.OUTPUT]) ,XIC(MC_CIP_AV01.CW.[CWD.OUTPUT]) OTE(MC_CIP_AV01_DR) ,XIC(S:FS) [OTU(MC_CIP_AV01.CW.[CWD.MANUAL]) ,LEQ(MC_CIP_AV01.CheckTime,0) MOV(Default_Check_Time,MC_CIP_AV01.CheckTime) ] ,[[XIC(MC_CIP_AV01_O) XIO(Item_Simulation_Flag) ,XIC(Item_Simulation_Flag) XIC(MC_CIP_AV01.CW.[CWD.OUTPUT]) XIO(MC_CIP_AV01.CW.[CWD.SIMFAIL]) ] OTE(MC_CIP_AV01.CW.[CWD.OPENFB]) ,[XIC(MC_CIP_AV01_C) XIO(Item_Simulation_Flag) ,XIC(Item_Simulation_Flag) XIO(MC_CIP_AV01.CW.[CWD.OUTPUT]) XIO(MC_CIP_AV01.CW.[CWD.SIMFAIL]) ] OTE(MC_CIP_AV01.CW.[CWD.CLOSEDFB]) ] ,[XIC(MC_CIP_AV01.CW.[CWD.OUTPUT]) XIO(MC_CIP_AV01.CW.[CWD.PREVSCAN]) ,XIO(MC_CIP_AV01.CW.[CWD.OUTPUT]) XIC(MC_CIP_AV01.CW.[CWD.PREVSCAN]) ] CLR(MC_CIP_AV01.CheckTimer) ,XIC(One_Second_One_Scan) LES(MC_CIP_AV01.CheckTimer,MC_CIP_AV01.CheckTime) ADD(MC_CIP_AV01.CheckTimer,1,MC_CIP_AV01.CheckTimer) ,XIO(MC_CIP_AV01.CW.[CWD.FAULT]) OTU(MC_CIP_AV01.CW.[CWD.FAULTLOGGED]) ,[GEQ(MC_CIP_AV01.CheckTimer,MC_CIP_AV01.CheckTime) [XIC(MC_CIP_AV01.CW.[CWD.OUTPUT]) [XIO(MC_CIP_AV01.CW.[CWD.OPENFB]) ,XIC(MC_CIP_AV01.CW.[CWD.CLOSEDFB]) ] ,XIO(MC_CIP_AV01.CW.[CWD.OUTPUT]) [XIC(MC_CIP_AV01.CW.[CWD.OPENFB]) ,XIO(MC_CIP_AV01.CW.[CWD.CLOSEDFB]) ] ] ,XIC(MC_CIP_AV01.CW.[CWD.FAULT]) XIC(Item_Faults_Are_Latched) ,XIC(MC_CIP_AV01.CW.[CWD.HIGHLIGHT]) ] XIO(MC_CIP_AV01.CW.[CWD.CHECKOFF]) XIO(Alarm_Reset) [OTE(MC_CIP_AV01.CW.[CWD.FAULT]) ,ALMD(MC_CIP_AV01_ALARM,0,0,0,0) ] ,XIC(MC_CIP_AV01.CW.[CWD.OUTPUT]) OTE(MC_CIP_AV01.CW.[CWD.PREVSCAN]) ];